// TIA Portal project "Despertador plclogiclab" (V16)

(* hardware
DEVICE "S7-1200 station_1"  S7-1200 Station
   slot 0: "Rack_0"  S7-1200 Rack  Rack  V1.0
   slot 1: "PLC_1"  CPU 1214C AC/DC/Rly  6ES7 214-1BG40-0XB0  V4.4
DEVICE "HMI_1"  TP2200 Comfort
   slot 0: "HMI_1"  TP2200 Comfort  6AV2 124-0XC02-0AX1  16.0.0.0
   slot 1: "HMI_RT_1"  TP2200 Comfort  6AV2 124-0XC02-0AX1  16.0.0.0
   slot 5: "HMI_1.IE_CP_1"  PROFINET Interface  16.0.0.0
      slot 1: "PROFINET Interface_1"  PROFINET Interface
         slot 1: "Port_1"  Port
         slot 2: "Port_2"  Port
   slot 6: "HMI_1.IE_CP_2"  PROFINET Interface  16.0.0.0
      slot 1: "PROFINET Interface_GBit"  PROFINET Interface
         slot 1: "Port_1"  Port
   slot 7: "HMI_1.MPI/DP_CP_1"  MPI/DP Interface  16.0.0.0
*)

// ===== PLC "PLC_1"  CPU 1214C AC/DC/Rly =====

VAR_GLOBAL   // PLC tag table "Default tag table"
   "stop_pb" AT %M3.1 : Bool;
   "start_pb" AT %M3.0 : Bool;
   "Tag_19" AT %I0.6 : Bool;
   "stop_alarm_pb" AT %M3.2 : Bool;
   "green pilot light" AT %Q0.0 : Bool;
   "Tag_9" AT %Q1.0 : Bool;
   "alarm" AT %Q0.7 : Bool;
   "lamp" AT %Q0.5 : Bool;
   "E. stop" AT %I0.0 : Bool;
   "System_Byte" AT %MB1 : Byte;
   "FirstScan" AT %M1.0 : Bool;
   "DiagStatusUpdate" AT %M1.1 : Bool;
   "AlwaysTRUE" AT %M1.2 : Bool;
   "AlwaysFALSE" AT %M1.3 : Bool;
   "DISABLE DEVICE" AT %M2.0 : Bool;
   "white_pilot_light" AT %Q0.2 : Bool;
END_VAR

DATA_BLOCK "alarma"   // DB1
{ S7_Optimized_Access := 'FALSE' }
VERSION : 0.1
   VAR
      horaactual : DTL;
      horaalarmainicio : DTL;
      horanuevai : DTL;
      stop : Bool;
      start : Bool;
      alarmaactivada : Bool;
      alarmasonando : Bool;
      status : Int;
      aux : Bool;
   END_VAR
BEGIN
END_DATA_BLOCK

// folder: System blocks/Program resources

DATA_BLOCK "timeralarma"   // DB2
{ S7_Optimized_Access := 'TRUE' }
AUTHOR : Simatic
FAMILY : IEC
NAME : IEC_TMR
VERSION : 1.0
// stored: InstanceOfName IEC_TIMER
"IEC_TIMER"
BEGIN
END_DATA_BLOCK

DATA_BLOCK "toff"   // DB3
{ S7_Optimized_Access := 'TRUE' }
AUTHOR : Simatic
FAMILY : IEC
NAME : IEC_TMR
VERSION : 1.0
// stored: InstanceOfName IEC_TIMER
"IEC_TIMER"
BEGIN
END_DATA_BLOCK

// folder: (top level)

ORGANIZATION_BLOCK "Main"   // OB1, LAD, ProgramCycle
TITLE = "Main Program Sweep (Cycle)"
{ S7_Optimized_Access := 'TRUE' }
VERSION : 0.1
// Alarma Diaria configurable para apagar un dispositivo por determinado tiempo
   VAR_INPUT
      Initial_Call : Bool;   // Initial call of this OB
      Remanence : Bool;   // =True, if remanent data are available
   END_VAR
   VAR_TEMP   // added for the SCL form of the ladder/FBD networks
      _w1 : Bool;
   END_VAR
BEGIN

REGION Network 1: start/stop system
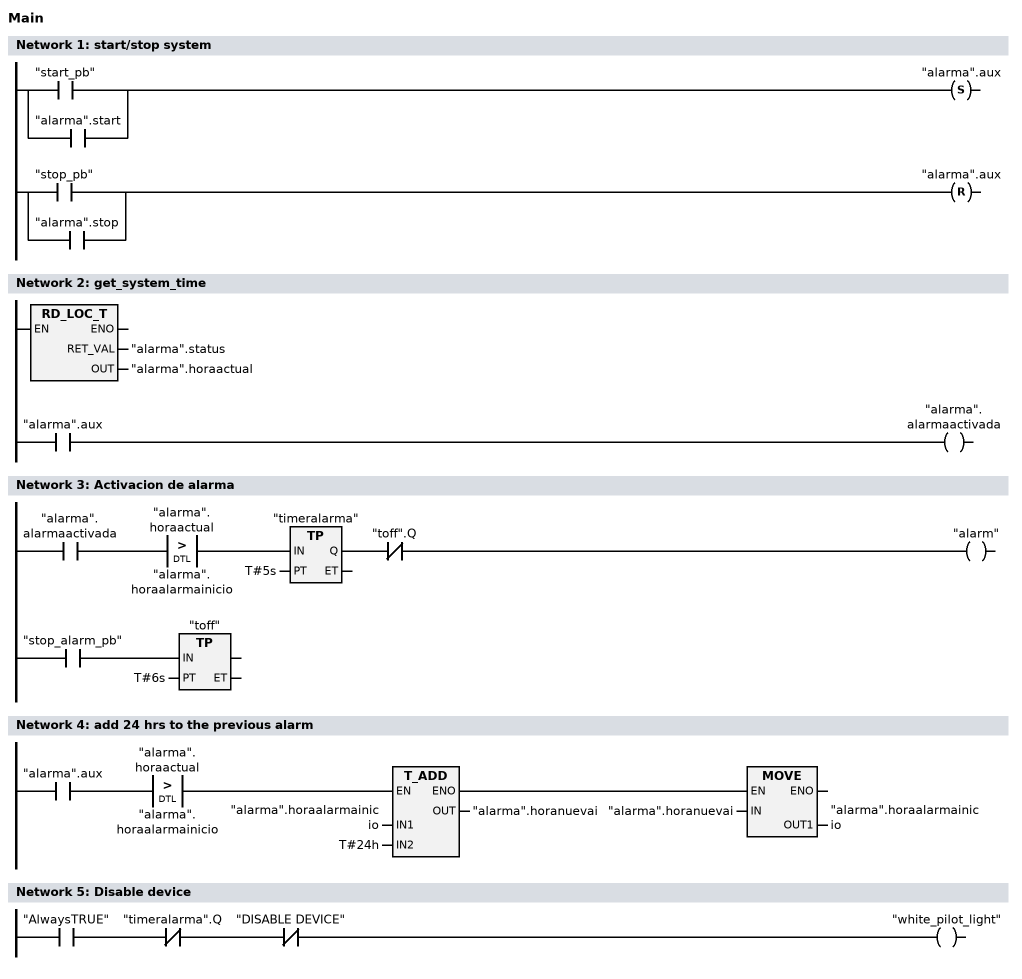
   RUNG wire#powerrail
      Contact( "start_pb" )
      wire#w1
      S_Coil( "alarma".aux )
   END_RUNG
   RUNG wire#powerrail
      Contact( "alarma".start )
   END_RUNG wire#w1
   RUNG wire#powerrail
      Contact( "stop_pb" )
      wire#w2
      R_Coil( "alarma".aux )
   END_RUNG
   RUNG wire#powerrail
      Contact( "alarma".stop )
   END_RUNG wire#w2
   // the same network as SCL:
   IF "start_pb" OR "alarma".start THEN "alarma".aux := TRUE; END_IF;
   IF "stop_pb" OR "alarma".stop THEN "alarma".aux := FALSE; END_IF;
END_REGION

REGION Network 2: get_system_time
   "alarma".status := RD_LOC_T(OUT => "alarma".horaactual);
   "alarma".alarmaactivada := "alarma".aux;
END_REGION

REGION Network 3: Activacion de alarma
   "timeralarma".TP(IN := "alarma".alarmaactivada AND ("alarma".horaactual > "alarma".horaalarmainicio),
                    PT := T#5s);
   "alarm" := "timeralarma".Q AND NOT "toff".Q;
   "toff".TP(IN := "stop_alarm_pb", PT := T#6s);
END_REGION

REGION Network 4: add 24 hrs to the previous alarm
   // ENO of a box is taken as its EN; it also drops when the box reports an error
   #_w1 := "alarma".aux AND ("alarma".horaactual > "alarma".horaalarmainicio);
   IF #_w1 THEN
       "alarma".horanuevai := T_ADD(IN1 := "alarma".horaalarmainicio, IN2 := T#24h);
       "alarma".horaalarmainicio := "alarma".horanuevai;
   END_IF;
END_REGION

REGION Network 5: Disable device
   RUNG wire#powerrail
      Contact( "AlwaysTRUE" )
      I_Contact( "timeralarma".Q )
      I_Contact( "DISABLE DEVICE" )
      Coil( "white_pilot_light" )
   END_RUNG
   // the same network as SCL:
   "white_pilot_light" := "AlwaysTRUE" AND NOT "timeralarma".Q AND NOT "DISABLE DEVICE";
END_REGION
END_ORGANIZATION_BLOCK

(* ===== HMI "HMI_RT_1" =====
system functions are stored by id; their names below are inferred from use
connection "HMI_Connection_1": ETHERNET, S7_1200_OMS

HMI tags "Default tag table"
   "alarma_horaactual" : DTL = PLC alarma.horaactual AT %DB1.DBX0.0, 100 ms
   "alarma_horaalarmainicio" : DTL = PLC alarma.horaalarmainicio AT %DB1.DBX12.0, 100 ms
   "Tag_16" : Bool = PLC lamp AT %Q0.5, 100 ms
   "alarma_start" : Bool = PLC alarma.start AT %DB1.DBX36.1, 100 ms
   "alarma_stop" : Bool = PLC alarma.stop AT %DB1.DBX36.0, 100 ms
   "DISABLE DEVICE" : Bool = PLC "DISABLE DEVICE" AT %M2.0, 100 ms
   "green pilot light" : Bool = PLC "green pilot light" AT %Q0.0, 100 ms
   "Tag_1" : Bool = PLC white_pilot_light AT %Q0.2, 100 ms
   "alarm" : Bool = PLC alarm AT %Q0.7, 100 ms

screen "Screen_1" 1920x1080
   GraphicView "Graphic view_1" at 0,0 size 1918x1076; Picture "Screenshot 2024-12-27 121323"
   Button "Button_1" at 774,680 size 390x136; TextOff 'ALARM CONFIG.'
      on Press: ActivateScreen("Screen_2", 0)
   TextField "Text field_1" at 824,172 size 382x91; Text 'WELCOME'

screen "Screen_2" 1920x1080
   GraphicView "Graphic view_1" at 0,3 size 1918x1076; Picture "Screenshot 2024-12-27 121323"
   Button "Button_1" at 832,734 size 303x86; TextOff 'MAIN'
      on Press: ActivateScreen("Screen_1", 0)
   IOField "I/O field_2" at 190,134 size 433x79; FormatPattern 9999999999999999999999999999999999999999
      ProcessValue <- "alarma_horaalarmainicio"
   IOField "I/O field_1" at 1343,134 size 429x79; FormatPattern 9999999999999999999999999999999999999999
      ProcessValue <- "alarma_horaactual"
   TextField "Text field_1" at 1526,224 size 102x47; Text 'TIME'
   TextField "Text field_2" at 324,220 size 197x43; Text 'ALARM SET'
   SymbolLibrary "Symbol library_1" at 370,278 size 279x160
   Button "Button_2" at 200,471 size 151x80; TextOff 'START'
      on Press: SetBit("alarma_start")
      on Release: ResetBit("alarma_start")
   Button "Button_3" at 645,469 size 151x80; TextOff 'STOP'
      on Press: SetBit("alarma_stop")
      on Release: ResetBit("alarma_stop")
   Rectangle "Rectangle_1" at 417,338 size 104x74
      Appearance <- "alarm"
   TextField "Text field_3" at 993,290 size 642x47; Text 'DISABLE DEVICE DURING ALARM'
   SymbolLibrary "Symbol library_2" at 1202,325 size 279x160
   Rectangle "Rectangle_2" at 1274,397 size 104x74
      Appearance <- "Tag_1"
   Switch "Switch_1" at 1139,523 size 304x136; CaptionText 'MANUAL SWITCH'; TextOff 'OFF'; TextOn 'ON'
      ProcessValue <- "DISABLE DEVICE"
*)